// TIA Portal project "DnomaidDBMS" (V13) (continued)
REGION Network 8: dA..Data Select
         L     #Network_8;
         T     #P_RET_VAL.MEM;
         A(;
         L     #COUNT.dA00;
         L     0;
         <>I;
         );
         A(;
         L     #COUNT.dA00;
         L     #QuantityDB;
         <=I;
         );
         JC    dA00;
         L     1;
         T     #COUNT.dA00;
         JU    dA00;
   dA00: NOP   0;
         L     #COUNT.dA00;
         JL    dAXX;
         JU    dAXX;
         JU    dA11;  //db[1]
         JU    dA21;  //db[2]
         JU    dA31;  //db[3]
         JU    dA41;  //db[4]
         JU    dA51;  //db[5]
         JU    dA61;  //db[6]
   dAXX: JU    dZFF;  //end
   dA11: NOP   0;
         L     #COUNT.dA00;
         T     #Status.Mem.SelctBBDDNum;
         SET;
         R     #AUX.FullDatabase;
         A     #Status.Perm.Push_nDB[1];
         AN    #Status.Mem.Full_nDB[1];
         =     #AUX.PushDatabase;
         JCN   dA12;
         L     #P_RET_VAL.MEM;
         T     #P_RET_VAL.V[1];
         T     #P_RET_VAL.V[2];
         CALL  FILL
         ( BVAL    := #ANY_DB1_FE,
           RET_VAL := #P_RET_VAL.V[1],
           BLK     := #ANY_DB1_IE
         );
         L     #P_RET_VAL.V[1];
         L     0;
         <>I;
         S     #FAULT;
         JC    END;
         CALL  FILL
         ( BVAL    := #IniData,
           RET_VAL := #P_RET_VAL.V[2],
           BLK     := #ANY_DB1_F
         );
         L     #P_RET_VAL.V[2];
         L     0;
         <>I;
         S     #FAULT;
         JC    END;
         R     #Status.Perm.Push_nDB[1];
         JU    dWFF;
   dA12: NOP   0;
         OPN   DB[ #LIST_DB_T.DbNumber[1]];
         LAR1  #""Address_104";
         L     LD[AR1, P#0.0];
         T     #AUX.LD_01;
         L     LW[AR1, P#4.0];
         T     #AUX.LW_01;
         L     LD[AR1, P#6.0];
         T     #AUX.LD_02;
         LAR1  #""Address_290";  //SEL
         L     #AUX.LD_01;
         T     LD[AR1, P#0.0];
         L     #AUX.LW_01;
         T     LW[AR1, P#4.0];
         L     #AUX.LD_02;
         T     LD[AR1, P#6.0];
         T     #P_ADR.I;
         LAR1  #""Address_113";
         L     LD[AR1, P#0.0];
         T     #AUX.LD_01;
         L     LW[AR1, P#4.0];
         T     #AUX.LW_01;
         L     LD[AR1, P#6.0];
         T     #AUX.LD_02;
         LAR1  #""Address_293";  //SEL
         L     #AUX.LD_01;
         T     LD[AR1, P#0.0];
         L     #AUX.LW_01;
         T     LW[AR1, P#4.0];
         L     #AUX.LD_02;
         T     LD[AR1, P#6.0];
         T     #P_ADR.F;
         JU    dAFF;
   dA21: NOP   0;
         L     #COUNT.dA00;
         T     #Status.Mem.SelctBBDDNum;
         SET;
         R     #AUX.FullDatabase;
         A     #Status.Perm.Push_nDB[2];
         AN    #Status.Mem.Full_nDB[2];
         =     #AUX.PushDatabase;
         JCN   dA22;
         L     #P_RET_VAL.MEM;
         T     #P_RET_VAL.V[1];
         T     #P_RET_VAL.V[2];
         CALL  FILL
         ( BVAL    := #ANY_DB2_FE,
           RET_VAL := #P_RET_VAL.V[1],
           BLK     := #ANY_DB2_IE
         );
         L     #P_RET_VAL.V[1];
         L     0;
         <>I;
         S     #FAULT;
         JC    END;
         CALL  FILL
         ( BVAL    := #IniData,
           RET_VAL := #P_RET_VAL.V[2],
           BLK     := #ANY_DB2_F
         );
         L     #P_RET_VAL.V[2];
         L     0;
         <>I;
         S     #FAULT;
         JC    END;
         R     #Status.Perm.Push_nDB[2];
         JU    dWFF;
   dA22: NOP   0;
         OPN   DB[ #LIST_DB_T.DbNumber[2]];
         LAR1  #""Address_119";
         L     LD[AR1, P#0.0];
         T     #AUX.LD_01;
         L     LW[AR1, P#4.0];
         T     #AUX.LW_01;
         L     LD[AR1, P#6.0];
         T     #AUX.LD_02;
         LAR1  #""Address_290";  //SEL
         L     #AUX.LD_01;
         T     LD[AR1, P#0.0];
         L     #AUX.LW_01;
         T     LW[AR1, P#4.0];
         L     #AUX.LD_02;
         T     LD[AR1, P#6.0];
         T     #P_ADR.I;
         LAR1  #""Address_126";
         L     LD[AR1, P#0.0];
         T     #AUX.LD_01;
         L     LW[AR1, P#4.0];
         T     #AUX.LW_01;
         L     LD[AR1, P#6.0];
         T     #AUX.LD_02;
         LAR1  #""Address_293";  //SELECT
         L     #AUX.LD_01;
         T     LD[AR1, P#0.0];
         L     #AUX.LW_01;
         T     LW[AR1, P#4.0];
         L     #AUX.LD_02;
         T     LD[AR1, P#6.0];
         T     #P_ADR.F;
         JU    dAFF;
   dA31: NOP   0;
         L     #COUNT.dA00;
         T     #Status.Mem.SelctBBDDNum;
         SET;
         R     #AUX.FullDatabase;
         A     #Status.Perm.Push_nDB[3];
         AN    #Status.Mem.Full_nDB[3];
         =     #AUX.PushDatabase;
         JCN   dA32;
         L     #P_RET_VAL.MEM;
         T     #P_RET_VAL.V[1];
         T     #P_RET_VAL.V[2];
         CALL  FILL
         ( BVAL    := #ANY_DB3_FE,
           RET_VAL := #P_RET_VAL.V[1],
           BLK     := #ANY_DB3_IE
         );
         L     #P_RET_VAL.V[1];
         L     0;
         <>I;
         S     #FAULT;
         JC    END;
         CALL  FILL
         ( BVAL    := #IniData,
           RET_VAL := #P_RET_VAL.V[2],
           BLK     := #ANY_DB3_F
         );
         L     #P_RET_VAL.V[2];
         L     0;
         <>I;
         S     #FAULT;
         JC    END;
         R     #Status.Perm.Push_nDB[3];
         JU    dWFF;
   dA32: NOP   0;
         OPN   DB[ #LIST_DB_T.DbNumber[3]];
         LAR1  #""Address_132";
         L     LD[AR1, P#0.0];
         T     #AUX.LD_01;
         L     LW[AR1, P#4.0];
         T     #AUX.LW_01;
         L     LD[AR1, P#6.0];
         T     #AUX.LD_02;
         LAR1  #""Address_290";  //SEL
         L     #AUX.LD_01;
         T     LD[AR1, P#0.0];
         L     #AUX.LW_01;
         T     LW[AR1, P#4.0];
         L     #AUX.LD_02;
         T     LD[AR1, P#6.0];
         T     #P_ADR.I;
         LAR1  #""Address_139";
         L     LD[AR1, P#0.0];
         T     #AUX.LD_01;
         L     LW[AR1, P#4.0];
         T     #AUX.LW_01;
         L     LD[AR1, P#6.0];
         T     #AUX.LD_02;
         LAR1  #""Address_293";  //SEL
         L     #AUX.LD_01;
         T     LD[AR1, P#0.0];
         L     #AUX.LW_01;
         T     LW[AR1, P#4.0];
         L     #AUX.LD_02;
         T     LD[AR1, P#6.0];
         T     #P_ADR.F;
         JU    dAFF;
   dA41: NOP   0;
         L     #COUNT.dA00;
         T     #Status.Mem.SelctBBDDNum;
         SET;
         R     #AUX.FullDatabase;
         A     #Status.Perm.Push_nDB[4];
         AN    #Status.Mem.Full_nDB[4];
         =     #AUX.PushDatabase;
         JCN   dA42;
         L     #P_RET_VAL.MEM;
         T     #P_RET_VAL.V[1];
         T     #P_RET_VAL.V[2];
         CALL  FILL
         ( BVAL    := #ANY_DB4_FE,
           RET_VAL := #P_RET_VAL.V[1],
           BLK     := #ANY_DB4_IE
         );
         L     #P_RET_VAL.V[1];
         L     0;
         <>I;
         S     #FAULT;
         JC    END;
         CALL  FILL
         ( BVAL    := #IniData,
           RET_VAL := #P_RET_VAL.V[2],
           BLK     := #ANY_DB4_F
         );
         L     #P_RET_VAL.V[2];
         L     0;
         <>I;
         S     #FAULT;
         JC    END;
         R     #Status.Perm.Push_nDB[4];
         JU    dWFF;
   dA42: NOP   0;
         OPN   DB[ #LIST_DB_T.DbNumber[4]];
         LAR1  #""Address_145";
         L     LD[AR1, P#0.0];
         T     #AUX.LD_01;
         L     LW[AR1, P#4.0];
         T     #AUX.LW_01;
         L     LD[AR1, P#6.0];
         T     #AUX.LD_02;
         LAR1  #""Address_290";  //SEL
         L     #AUX.LD_01;
         T     LD[AR1, P#0.0];
         L     #AUX.LW_01;
         T     LW[AR1, P#4.0];
         L     #AUX.LD_02;
         T     LD[AR1, P#6.0];
         T     #P_ADR.I;
         LAR1  #""Address_152";
         L     LD[AR1, P#0.0];
         T     #AUX.LD_01;
         L     LW[AR1, P#4.0];
         T     #AUX.LW_01;
         L     LD[AR1, P#6.0];
         T     #AUX.LD_02;
         LAR1  #""Address_293";  //SEL
         L     #AUX.LD_01;
         T     LD[AR1, P#0.0];
         L     #AUX.LW_01;
         T     LW[AR1, P#4.0];
         L     #AUX.LD_02;
         T     LD[AR1, P#6.0];
         T     #P_ADR.F;
         JU    dAFF;
   dA51: NOP   0;
         L     #COUNT.dA00;
         T     #Status.Mem.SelctBBDDNum;
         SET;
         R     #AUX.FullDatabase;
         A     #Status.Perm.Push_nDB[5];
         AN    #Status.Mem.Full_nDB[5];
         =     #AUX.PushDatabase;
         JCN   dA52;
         L     #P_RET_VAL.MEM;
         T     #P_RET_VAL.V[1];
         T     #P_RET_VAL.V[2];
         CALL  FILL
         ( BVAL    := #ANY_DB5_FE,
           RET_VAL := #P_RET_VAL.V[1],
           BLK     := #ANY_DB5_IE
         );
         L     #P_RET_VAL.V[1];
         L     0;
         <>I;
         S     #FAULT;
         JC    END;
         CALL  FILL
         ( BVAL    := #IniData,
           RET_VAL := #P_RET_VAL.V[2],
           BLK     := #ANY_DB5_F
         );
         L     #P_RET_VAL.V[2];
         L     0;
         <>I;
         S     #FAULT;
         JC    END;
         R     #Status.Perm.Push_nDB[5];
         JU    dWFF;
   dA52: NOP   0;
         OPN   DB[ #LIST_DB_T.DbNumber[5]];
         LAR1  #""Address_158";
         L     LD[AR1, P#0.0];
         T     #AUX.LD_01;
         L     LW[AR1, P#4.0];
         T     #AUX.LW_01;
         L     LD[AR1, P#6.0];
         T     #AUX.LD_02;
         LAR1  #""Address_290";  //SEL
         L     #AUX.LD_01;
         T     LD[AR1, P#0.0];
         L     #AUX.LW_01;
         T     LW[AR1, P#4.0];
         L     #AUX.LD_02;
         T     LD[AR1, P#6.0];
         T     #P_ADR.I;
         LAR1  #""Address_165";
         L     LD[AR1, P#0.0];
         T     #AUX.LD_01;
         L     LW[AR1, P#4.0];
         T     #AUX.LW_01;
         L     LD[AR1, P#6.0];
         T     #AUX.LD_02;
         LAR1  #""Address_293";  //SEL
         L     #AUX.LD_01;
         T     LD[AR1, P#0.0];
         L     #AUX.LW_01;
         T     LW[AR1, P#4.0];
         L     #AUX.LD_02;
         T     LD[AR1, P#6.0];
         T     #P_ADR.F;
         JU    dAFF;
   dA61: NOP   0;
         L     #COUNT.dA00;
         T     #Status.Mem.SelctBBDDNum;
         SET;
         R     #AUX.FullDatabase;
         A     #Status.Perm.Push_nDB[6];
         AN    #Status.Mem.Full_nDB[6];
         =     #AUX.PushDatabase;
         JCN   dA62;
         L     #P_RET_VAL.MEM;
         T     #P_RET_VAL.V[1];
         T     #P_RET_VAL.V[2];
         CALL  FILL
         ( BVAL    := #ANY_DB6_FE,
           RET_VAL := #P_RET_VAL.V[1],
           BLK     := #ANY_DB6_IE
         );
         L     #P_RET_VAL.V[1];
         L     0;
         <>I;
         S     #FAULT;
         JC    END;
         CALL  FILL
         ( BVAL    := #IniData,
           RET_VAL := #P_RET_VAL.V[2],
           BLK     := #ANY_DB6_F
         );
         L     #P_RET_VAL.V[2];
         L     0;
         <>I;
         S     #FAULT;
         JC    END;
         R     #Status.Perm.Push_nDB[6];
         JU    dWFF;
   dA62: NOP   0;
         OPN   DB[ #LIST_DB_T.DbNumber[6]];
         LAR1  #""Address_171";
         L     LD[AR1, P#0.0];
         T     #AUX.LD_01;
         L     LW[AR1, P#4.0];
         T     #AUX.LW_01;
         L     LD[AR1, P#6.0];
         T     #AUX.LD_02;
         LAR1  #""Address_290";  //SEL
         L     #AUX.LD_01;
         T     LD[AR1, P#0.0];
         L     #AUX.LW_01;
         T     LW[AR1, P#4.0];
         L     #AUX.LD_02;
         T     LD[AR1, P#6.0];
         T     #P_ADR.I;
         LAR1  #""Address_178";
         L     LD[AR1, P#0.0];
         T     #AUX.LD_01;
         L     LW[AR1, P#4.0];
         T     #AUX.LW_01;
         L     LD[AR1, P#6.0];
         T     #AUX.LD_02;
         LAR1  #""Address_293";  //SEL
         L     #AUX.LD_01;
         T     LD[AR1, P#0.0];
         L     #AUX.LW_01;
         T     LW[AR1, P#4.0];
         L     #AUX.LD_02;
         T     LD[AR1, P#6.0];
         T     #P_ADR.F;
         JU    dAFF;
   dAFF: NOP   0;
END_REGION

REGION Network 9: dC..Data Search empty space
         LAR1  #P_ADR.I;
         JU    dC00;
   dC00: NOP   0;
         L     #Network_9;
         T     #P_RET_VAL.MEM;
         TAR1;
         T     #SAVE_AR1.dC00;
         L     1;
   dC01: NOP   0;
         T     #COUNT.dC00;
         L     DBB[AR1, P#0.0];
         L     ' ';
         <>I;
         =     #AUX.DifferentValue;
         AN    #AUX.DifferentValue;
         JC    dCFF;
         L     #P_ADR.F;
         L     #SAVE_AR1.dC00;
         <=D;
         =     #AUX.FullDatabase;
         A     #AUX.FullDatabase;
         JC    dCWF;
         L     P#1.0;
         +AR1;
         L     #COUNT.dC00;
         LOOP  dC01;
         L     #SAVE_AR1.dC00;
         LAR1;
         L     #LENGTH.PointerData;
         +AR1;
         JU    dC00;
END_REGION

REGION Network 10: dC..Data Full
         JU    dCWF;
   dCWF: NOP   0;
         L     #Network_10;
         T     #P_RET_VAL.MEM;
         AN    #AUX.FullDatabase;
         JC    dCWW;
         L     #Status.Mem.SelctBBDDNum;
         JL    dCXX;
         JU    dCEE;  //fault
         JU    dC11;  //db[1]
         JU    dC12;  //db[2]
         JU    dC13;  //db[3]
         JU    dC14;  //db[4]
         JU    dC15;  //db[5]
         JU    dC16;  //db[6]
   dCXX: JU    dCEE;  //fault
   dC11: NOP   0;
         A     #AUX.FullDatabase;
         =     #Status.Mem.Full_nDB[1];
         JU    dCWW;
   dC12: NOP   0;
         A     #AUX.FullDatabase;
         =     #Status.Mem.Full_nDB[2];
         JU    dCWW;
   dC13: NOP   0;
         A     #AUX.FullDatabase;
         =     #Status.Mem.Full_nDB[3];
         JU    dCWW;
   dC14: NOP   0;
         A     #AUX.FullDatabase;
         =     #Status.Mem.Full_nDB[4];
         JU    dCWW;
   dC15: NOP   0;
         A     #AUX.FullDatabase;
         =     #Status.Mem.Full_nDB[5];
         JU    dCWW;
   dC16: NOP   0;
         A     #AUX.FullDatabase;
         =     #Status.Mem.Full_nDB[6];
         JU    dCWW;
   dCEE: NOP   0;
         SET;
         S     #FAULT;
         JU    END;
   dCWW: NOP   0;
         JU    dWFF;
         JU    dCFF;
   dCFF: NOP   0;
END_REGION

REGION Network 11: dD..Data Find space
         JU    dD00;
   dD00: NOP   0;
         L     #Network_11;
         T     #P_RET_VAL.MEM;
         L     #SAVE_AR1.dC00;
         LAR1;
         L     #LENGTH.PointerData;
         +AR1;
         L     #P_ADR.F;
         TAR1;
         <D;
         JC    dWFF;
         JU    dDFF;
   dDFF: NOP   0;
END_REGION

REGION Network 12: dE..Data Find data
         JU    dE00;
   dE00: NOP   0;
         L     #Network_12;
         T     #P_RET_VAL.MEM;
         TAR1;
         T     #SAVE_AR1.dE00;
         L     1;
   dE01: NOP   0;
         T     #COUNT.dE00;
         L     DBB[AR1, P#0.0];
         L     ' ';
         ==I;
         =     #AUX.EmptyData;
         AN    #AUX.EmptyData;
         JC    dEFF;
         L     #P_ADR.F;
         L     #SAVE_AR1.dE00;
         <=D;
         JC    dWFF;
         L     P#1.0;
         +AR1;
         L     #COUNT.dE00;
         LOOP  dE01;
         L     #SAVE_AR1.dE00;
         LAR1;
         L     #LENGTH.PointerData;
         +AR1;
         JU    dE00;
         JU    dEFF;
   dEFF: NOP   0;
END_REGION

REGION Network 13: dF..Data Move data
         JU    dF01;
   dF01: NOP   0;
         L     #Network_13;
         T     #P_RET_VAL.MEM;
         L     #SAVE_AR1.dE00;
         T     #P_ADR.F;
         LAR1  #""Address_293";
         T     LD[AR1, P#6.0];
         L     #SAVE_AR1.dC00;
         T     #P_ADR.I;
         LAR1  #""Address_290";
         T     LD[AR1, P#6.0];
         LAR1;
         L     #P_RET_VAL.MEM;
         T     #P_RET_VAL.V[1];
         T     #P_RET_VAL.V[2];
         CALL  FILL
         ( BVAL    := #ANY_DB_SELECT_F,
           RET_VAL := #P_RET_VAL.V[1],
           BLK     := #ANY_DB_SELECT_I
         );
         L     #P_RET_VAL.V[1];
         L     0;
         <>I;
         S     #FAULT;
         JC    END;
         CALL  FILL
         ( BVAL    := #IniData,
           RET_VAL := #P_RET_VAL.V[2],
           BLK     := #ANY_DB_SELECT_F
         );
         L     #P_RET_VAL.V[2];
         L     0;
         <>I;
         S     #FAULT;
         JC    END;
         JU    dZFF;
   dWFF: NOP   0;
         L     #COUNT.dA00;
         +     1;
         T     #COUNT.dA00;
         L     #QuantityDB;
         >I;
         JC    dZFF;
         JU    dA00;
   //--->END
         JU    dZFF;
   dZFF: NOP   0;
END_REGION

REGION Network 14: fA..Query
         JU    fA0X;
   fA0X: NOP   0;
         L     #Network_14;
         T     #P_RET_VAL.MEM;
         AN    #Request.Query.Request;
         R     #Response.Query.DataAvailable;
         R     #Response.Query.DataNotAvailable;
         NOT;
         FP    #FP_REQUEST.QueryDB;
         JC    fA0Y;
         JU    fBFF;
   fA0Y: NOP   0;
         L     #P_RET_VAL.MEM;
         T     #P_RET_VAL.V[1];
         T     #P_RET_VAL.V[2];
         CALL  FILL
         ( BVAL    := #Request.Query.BarcodeDig,
           RET_VAL := #P_RET_VAL.V[1],
           BLK     := #DigitFilter
         );
         L     #P_RET_VAL.V[1];
         L     0;
         <>I;
         S     #FAULT;
         JC    END;
         JU    jA00;  //Goto Data input filters
   fAR2: NOP   0;  //Return Data input filters
         CALL  FILL
         ( BVAL    := #DigitFilter,
           RET_VAL := #P_RET_VAL.V[2],
           BLK     := #QueryData
         );
         L     #P_RET_VAL.V[2];
         L     0;
         <>I;
         S     #FAULT;
         JC    END;
         CALL  FILL
         ( BVAL    := #IniData,
           RET_VAL := #P_RET_VAL.V[3],
           BLK     := #Response.QueryDataAvailable
         );
         L     #P_RET_VAL.V[3];
         L     0;
         <>I;
         S     #FAULT;
         JC    END;
         AN    #DataInputOK;
         JC    fB50;  //Error data input
         L     1;
         T     #COUNT.fA00;
   fA00: NOP   0;
         L     #COUNT.fA00;
         JL    fAXX;
         JU    fAXX;
         JU    fA11;  //db[1]
         JU    fA21;  //db[2]
         JU    fA31;  //db[3]
         JU    fA41;  //db[4]
         JU    fA51;  //db[5]
         JU    fA61;  //db[6]
         JU    fB40;  //end
   fAXX: JU    fAEE;  //fault
   fA11: NOP   0;
         OPN   DB[ #LIST_DB_T.DbNumber[1]];
         LAR1  #P_ADR.I_DB[1];
         L     #NumDataArrayDB[1];
         JU    fA10;
   fA21: NOP   0;
         OPN   DB[ #LIST_DB_T.DbNumber[2]];
         LAR1  #P_ADR.I_DB[2];
         L     #NumDataArrayDB[2];
         JU    fA10;
   fA31: NOP   0;
         OPN   DB[ #LIST_DB_T.DbNumber[3]];
         LAR1  #P_ADR.I_DB[3];
         L     #NumDataArrayDB[3];
         JU    fA10;
   fA41: NOP   0;
         OPN   DB[ #LIST_DB_T.DbNumber[4]];
         LAR1  #P_ADR.I_DB[4];
         L     #NumDataArrayDB[4];
         JU    fA10;
   fA51: NOP   0;
         OPN   DB[ #LIST_DB_T.DbNumber[5]];
         LAR1  #P_ADR.I_DB[5];
         L     #NumDataArrayDB[5];
         JU    fA10;
   fA61: NOP   0;
         OPN   DB[ #LIST_DB_T.DbNumber[6]];
         LAR1  #P_ADR.I_DB[6];
         L     #NumDataArrayDB[6];
         JU    fA10;
   fA10: NOP   0;
         T     #COUNT.fA01;
         TAR1;
         T     #SAVE_AR1.fA10;
         SET;
   //-------------------------------
         TAR1;
         T     #P_ADR.SAVE_COMP_01;
         T     #P_ADR.COMP_01;
         L     #""Address_347";
         T     #P_ADR.COMP_02;
         SET;
         R     #AUX.DifferentValue;
         L     #LENGTH.Code;
   fMP0: NOP   0;
         T     #COUNT.fA02;
         LAR1  #P_ADR.COMP_01;
         L     DBB[AR1, P#0.0];
         LAR1  #P_ADR.COMP_02;
         L     DIB[AR1, P#0.0];
         <>I;
         S     #AUX.DifferentValue;
         L     P#1.0;
         L     #P_ADR.COMP_01;
         +D;
         T     #P_ADR.COMP_01;
         L     P#1.0;
         L     #P_ADR.COMP_02;
         +D;
         T     #P_ADR.COMP_02;
         L     #COUNT.fA02;
         LOOP  fMP0;
         LAR1  #P_ADR.SAVE_COMP_01;
   //-------------------------------
         AN    #AUX.DifferentValue;
         JC    fB20;
         L     #LENGTH.PointerData;
         +AR1;
         L     #COUNT.fA01;
         LOOP  fA10;
         JU    fWFF;
   fWFF: NOP   0;
         L     #COUNT.fA00;
         +     1;
         T     #COUNT.fA00;
         L     #QuantityDB;
         >I;
         JC    fB40;
         JU    fA00;
   fAEE: NOP   0;
         SET;
         S     #FAULT;
         JU    END;
         JU    fAFF;
   fAFF: NOP   0;
         JU    END;
   fB20: NOP   0;
         L     #COUNT.fA00;
         JL    fB3X;
         JU    fB3X;
         JU    fB31;  //db[1]
         JU    fB32;  //db[2]
         JU    fB33;  //db[3]
         JU    fB34;  //db[4]
         JU    fB35;  //db[5]
         JU    fB36;  //db[6]
   fB3X: JU    fB3E;  //fault
   fB31: NOP   0;
         LAR1  #""Address_104";
         JU    fB3F;
   fB32: NOP   0;
         LAR1  #""Address_119";
         JU    fB3F;
   fB33: NOP   0;
         LAR1  #""Address_132";
         JU    fB3F;
   fB34: NOP   0;
         LAR1  #""Address_145";
         JU    fB3F;
   fB35: NOP   0;
         LAR1  #""Address_158";
         JU    fB3F;
   fB36: NOP   0;
         LAR1  #""Address_171";
         JU    fB3F;
   fB3E: NOP   0;
         SET;
         S     #FAULT;
         JU    END;
         JU    fB3F;
   fB3F: NOP   0;
         L     LD[AR1, P#0.0];
         T     #AUX.LD_01;
         L     LW[AR1, P#4.0];
         T     #AUX.LW_01;
         T     #PAUXnDB;
         LAR1  #""Address_381";
         L     #AUX.LD_01;
         T     LD[AR1, P#0.0];
         L     #AUX.LW_01;
         T     LW[AR1, P#4.0];
         L     #SAVE_AR1.fA10;
         T     LD[AR1, P#6.0];
         L     #P_RET_VAL.MEM;
         T     #P_RET_VAL.V[1];
         CALL  FILL
         ( BVAL    := #ANY_DB_QUERY,
           RET_VAL := #P_RET_VAL.V[1],
           BLK     := #Response.QueryDataAvailable
         );
         L     #P_RET_VAL.V[1];
         L     0;
         <>I;
         S     #FAULT;
         JC    END;
         S     #Response.Query.DataAvailable;
         R     #Response.Query.DataNotAvailable;
         L     #LogDataAvailable;
         T     #Log.Request;
         JU    fB50;
   fB40: NOP   0;
         SET;
         R     #Response.Query.DataAvailable;
         S     #Response.Query.DataNotAvailable;
         L     #LogDataNotAvailable;
         T     #Log.Request;
   fB50: NOP   0;
         A     #DataInputOK;
         JC    fB51;  //Error data input
         L     #LogDataInputNOK;
         T     #Log.Request;
   fB51: NOP   0;
         L     #P_RET_VAL.MEM;
         T     #P_RET_VAL.V[1];
         CALL  FILL
         ( BVAL    := #QueryData,
           RET_VAL := #P_RET_VAL.V[1],
           BLK     := #Response.Query.BarcodeDig
         );
         L     #P_RET_VAL.V[1];
         L     0;
         <>I;
         S     #FAULT;
         JC    END;
         CALL  FILL
         ( BVAL    := #QueryData,
           RET_VAL := #P_RET_VAL.V[2],
           BLK     := #Log.DatabaseTable
         );
         L     #P_RET_VAL.V[2];
         L     0;
         <>I;
         S     #FAULT;
         JC    END;
         CALL  FILL
         ( BVAL    := #DateTime,
           RET_VAL := #P_RET_VAL.V[3],
           BLK     := #Log.DatabaseTable.DateTime
         );
         L     #P_RET_VAL.V[3];
         L     0;
         <>I;
         S     #FAULT;
         JC    END;
         JU    fBFF;
   fBFF: NOP   0;
END_REGION

REGION Network 15: gA..Insert
         JU    gA00;
   gA00: NOP   0;
         L     #Network_15;
         T     #P_RET_VAL.MEM;
         SET;
   //      R     #AUX.StatusPermInsert_nDB
         AN    #Request.Insert.Request;
         R     #Response.Insert.Completed;
         L     #QuantityDB;
         T     #COUNT.gA00;
         NOP   0;
         SET;
         L     #COUNT.gA00;
         JL    gAXX;
         JU    gAXX;
         JU    gA11;  //db[1]
         JU    gA21;  //db[2]
         JU    gA31;  //db[3]
         JU    gA41;  //db[4]
         JU    gA51;  //db[5]
         JU    gA61;  //db[6]
   gAXX: JU    gAEE;  //fault
   gA11: NOP   0;
         A     #Status.Perm.Insert_nDB[1];
         JU    gA01;
   gA21: NOP   0;
         A     #Status.Perm.Insert_nDB[2];
         JU    gA01;
   gA31: NOP   0;
         A     #Status.Perm.Insert_nDB[3];
         JU    gA01;
   gA41: NOP   0;
         A     #Status.Perm.Insert_nDB[4];
         JU    gA01;
   gA51: NOP   0;
         A     #Status.Perm.Insert_nDB[5];
         JU    gA01;
   gA61: NOP   0;
         A     #Status.Perm.Insert_nDB[6];
         JU    gA01;
   gAEE: NOP   0;
         SET;
         S     #FAULT;
         JU    END;
   gA01: NOP   0;
         =     #AUX.StatusPermInsert_nDB;
         A     #AUX.TON_StatusPermInsert_nDB;
         AN    #Status.Mem.FillAll;
         AN    #Status.Fb_Fault;
         =     #Status.Perm.Insert;
         A     #FULL;  //Data base full
         JC    gA02;
         A     #Request.Query.Request;
         JC    gAFF;
         A     #AUX.TON_StatusPermInsert_nDB;
   gA02: NOP   0;
         A     #Request.Insert.Request;
         FP    #FP_REQUEST.InsertDB;
         JC    gA03;
         JU    gAFF;
   gA03: NOP   0;
         L     #P_RET_VAL.MEM;
         T     #P_RET_VAL.V[1];
         T     #P_RET_VAL.V[2];
         T     #P_RET_VAL.V[3];
         T     #P_RET_VAL.V[4];
         T     #P_RET_VAL.V[5];
         CALL  FILL
         ( BVAL    := #Request.Insert.BarcodeData,
           RET_VAL := #P_RET_VAL.V[1],
           BLK     := #DigitFilter
         );
         L     #P_RET_VAL.V[1];
         L     0;
         <>I;
         S     #FAULT;
         JC    END;
         JU    jA00;  //Goto Data input filters
   gAR2: NOP   0;  //Return Data input filters
         CALL  FILL
         ( BVAL    := #DigitFilter,
           RET_VAL := #P_RET_VAL.V[2],
           BLK     := #InsertData.BarcodeData
         );
         L     #P_RET_VAL.V[2];
         L     0;
         <>I;
         S     #FAULT;
         JC    END;
         CALL  FILL
         ( BVAL    := #DateTime,
           RET_VAL := #P_RET_VAL.V[3],
           BLK     := #InsertData.DateTime
         );
         L     #P_RET_VAL.V[3];
         L     0;
         <>I;
         S     #FAULT;
         JC    END;
         AN    #DataInputOK;
         S     #DATA_ERROR;
         JC    gA05;  //Error data input
         A     #FULL;
         S     #DATA_ERROR;
         JC    gA06;  //Data base full
         L     #COUNT.gA00;
         JL    gBXX;
         JU    gBXX;
         JU    gB11;  //db[1]
         JU    gB21;  //db[2]
         JU    gB31;  //db[3]
         JU    gB41;  //db[4]
         JU    gB51;  //db[5]
         JU    gB61;  //db[6]
   gBXX: JU    gBEE;  //fault
   gB11: NOP   0;
         CALL  FILL
         ( BVAL    := #InsertData,
           RET_VAL := #P_RET_VAL.V[3],
           BLK     := #ANY_DB1_F
         );
         L     #P_RET_VAL.V[3];
         L     0;
         <>I;
         S     #FAULT;
         JC    END;
         JU    gA04;
   gB21: NOP   0;
         CALL  FILL
         ( BVAL    := #InsertData,
           RET_VAL := #P_RET_VAL.V[3],
           BLK     := #ANY_DB2_F
         );
         L     #P_RET_VAL.V[3];
         L     0;
         <>I;
         S     #FAULT;
         JC    END;
         JU    gA04;
   gB31: NOP   0;
         CALL  FILL
         ( BVAL    := #InsertData,
           RET_VAL := #P_RET_VAL.V[3],
           BLK     := #ANY_DB3_F
         );
         L     #P_RET_VAL.V[3];
         L     0;
         <>I;
         S     #FAULT;
         JC    END;
         JU    gA04;
   gB41: NOP   0;
         CALL  FILL
         ( BVAL    := #InsertData,
           RET_VAL := #P_RET_VAL.V[3],
           BLK     := #ANY_DB4_F
         );
         L     #P_RET_VAL.V[3];
         L     0;
         <>I;
         S     #FAULT;
         JC    END;
         JU    gA04;
   gB51: NOP   0;
         CALL  FILL
         ( BVAL    := #InsertData,
           RET_VAL := #P_RET_VAL.V[3],
           BLK     := #ANY_DB5_F
         );
         L     #P_RET_VAL.V[3];
         L     0;
         <>I;
         S     #FAULT;
         JC    END;
         JU    gA04;
   gB61: NOP   0;
         CALL  FILL
         ( BVAL    := #InsertData,
           RET_VAL := #P_RET_VAL.V[3],
           BLK     := #ANY_DB6_F
         );
         L     #P_RET_VAL.V[3];
         L     0;
         <>I;
         S     #FAULT;
         JC    END;
         JU    gA04;
   gBEE: NOP   0;
         SET;
         S     #FAULT;
         JU    END;
   gA04: NOP   0;
         CALL  FILL
         ( BVAL    := #InsertData,
           RET_VAL := #P_RET_VAL.V[4],
           BLK     := #Response.InsertData
         );
         L     #P_RET_VAL.V[4];
         L     0;
         <>I;
         S     #FAULT;
         JC    END;
         S     #Response.Insert.Completed;
         L     #LogInsert;
         T     #Log.Request;
         A     #DataInputOK;
         JC    gA07;
   gA05: NOP   0;
         L     #LogDataInputNOK;  //Data input NOK
         T     #Log.Request;
         SET;
         JU    gA07;
   gA06: NOP   0;
         L     #LogFullData;  //Data base full
         T     #Log.Request;
         SET;
         JU    gA07;
   gA07: NOP   0;
         CALL  FILL
         ( BVAL    := #InsertData,
           RET_VAL := #P_RET_VAL.V[5],
           BLK     := #Log.DatabaseTable
         );
         L     #P_RET_VAL.V[5];
         L     0;
         <>I;
         S     #FAULT;
         JC    END;
         JU    gAFF;
   gAFF: NOP   0;
END_REGION

REGION Network 16: hA..Delete
         JU    hA0X;
   hA0X: NOP   0;
         L     #Network_16;
         T     #P_RET_VAL.MEM;
         AN    #Request.Delete.Request;
         R     #Response.Delete.Completed;
         NOT;
         FP    #FP_REQUEST.DeleteDB;
         JC    hA0Y;
         JU    hBFF;
   hA0Y: NOP   0;
         L     #P_RET_VAL.MEM;
         T     #P_RET_VAL.V[1];
         T     #P_RET_VAL.V[2];
         CALL  FILL
         ( BVAL    := #Request.Delete.BarcodeDig,
           RET_VAL := #P_RET_VAL.V[1],
           BLK     := #DigitFilter
         );
         L     #P_RET_VAL.V[1];
         L     0;
         <>I;
         S     #FAULT;
         JC    END;
         JU    jA00;  //Goto Data input filters
   hAR2: NOP   0;  //Return Data input filters
         CALL  FILL
         ( BVAL    := #DigitFilter,
           RET_VAL := #P_RET_VAL.V[2],
           BLK     := #DeleteData
         );
         L     #P_RET_VAL.V[2];
         L     0;
         <>I;
         S     #FAULT;
         JC    END;
         CALL  FILL
         ( BVAL    := #IniData,
           RET_VAL := #P_RET_VAL.V[3],
           BLK     := #Response.DeleteData
         );
         L     #P_RET_VAL.V[3];
         L     0;
         <>I;
         S     #FAULT;
         AN    #DataInputOK;
         JC    hB3G;  //Error data input
         L     1;
         T     #COUNT.hA00;
   hA00: NOP   0;
         L     #COUNT.hA00;
         JL    hAXX;
         JU    hAXX;
         JU    hA11;  //db[1]
         JU    hA21;  //db[2]
         JU    hA31;  //db[3]
         JU    hA41;  //db[4]
         JU    hA51;  //db[5]
         JU    hA61;  //db[6]
         JU    hB40;  //end
   hAXX: JU    hAEE;  //fault
   hA11: NOP   0;
         OPN   DB[ #LIST_DB_T.DbNumber[1]];
         LAR1  #P_ADR.I_DB[1];
         L     #NumDataArrayDB[1];
         JU    hA10;
   hA21: NOP   0;
         OPN   DB[ #LIST_DB_T.DbNumber[2]];
         LAR1  #P_ADR.I_DB[2];
         L     #NumDataArrayDB[2];
         JU    hA10;
   hA31: NOP   0;
         OPN   DB[ #LIST_DB_T.DbNumber[3]];
         LAR1  #P_ADR.I_DB[3];
         L     #NumDataArrayDB[3];
         JU    hA10;
   hA41: NOP   0;
         OPN   DB[ #LIST_DB_T.DbNumber[4]];
         LAR1  #P_ADR.I_DB[4];
         L     #NumDataArrayDB[4];
         JU    hA10;
   hA51: NOP   0;
         OPN   DB[ #LIST_DB_T.DbNumber[5]];
         LAR1  #P_ADR.I_DB[5];
         L     #NumDataArrayDB[5];
         JU    hA10;
   hA61: NOP   0;
         OPN   DB[ #LIST_DB_T.DbNumber[6]];
         LAR1  #P_ADR.I_DB[6];
         L     #NumDataArrayDB[6];
         JU    hA10;
   hA10: NOP   0;
         T     #COUNT.hA01;
         TAR1;
         T     #SAVE_AR1.hA10;
         SET;
   //-------------------------------
         TAR1;
         T     #P_ADR.SAVE_COMP_01;
         T     #P_ADR.COMP_01;
         L     #""Address_433";
         T     #P_ADR.COMP_02;
         SET;
         R     #AUX.DifferentValue;
         L     #LENGTH.Code;
   hMP0: NOP   0;
         T     #COUNT.hA02;
         LAR1  #P_ADR.COMP_01;
         L     DBB[AR1, P#0.0];
         LAR1  #P_ADR.COMP_02;
         L     DIB[AR1, P#0.0];
         <>I;
         S     #AUX.DifferentValue;
         L     P#1.0;
         L     #P_ADR.COMP_01;
         +D;
         T     #P_ADR.COMP_01;
         L     P#1.0;
         L     #P_ADR.COMP_02;
         +D;
         T     #P_ADR.COMP_02;
         L     #COUNT.hA02;
         LOOP  hMP0;
         LAR1  #P_ADR.SAVE_COMP_01;
   //-------------------------------
         AN    #AUX.DifferentValue;
         JC    hB20;
         L     #LENGTH.PointerData;
         +AR1;
         L     #COUNT.hA01;
         LOOP  hA10;
         JU    hWFF;
   hWFF: NOP   0;
         L     #COUNT.hA00;
         +     1;
         T     #COUNT.hA00;
         L     #QuantityDB;
         >I;
         JC    hB40;
         JU    hA00;
   hAEE: NOP   0;
         SET;
         S     #FAULT;
         JU    END;
         JU    hAFF;
   hAFF: NOP   0;
         JU    END;
   hB20: NOP   0;
         NOP   0;
         L     #COUNT.hA00;
         JL    hB3X;
         JU    hB3X;
         JU    hB31;  //db[1]
         JU    hB32;  //db[2]
         JU    hB33;  //db[3]
         JU    hB34;  //db[4]
         JU    hB35;  //db[5]
         JU    hB36;  //db[6]
   hB3X: JU    hB3E;  //fault
   hB31: NOP   0;
         LAR1  #""Address_104";
         JU    hB3F;
   hB32: NOP   0;
         LAR1  #""Address_119";
         JU    hB3F;
   hB33: NOP   0;
         LAR1  #""Address_132";
         JU    hB3F;
   hB34: NOP   0;
         LAR1  #""Address_145";
         JU    hB3F;
   hB35: NOP   0;
         LAR1  #""Address_158";
         JU    hB3F;
   hB36: NOP   0;
         LAR1  #""Address_171";
         JU    hB3F;
   hB3E: NOP   0;
         SET;
         S     #FAULT;
         JU    END;
         JU    hB3F;
   hB3F: NOP   0;
         L     LD[AR1, P#0.0];
         T     #AUX.LD_01;
         L     LW[AR1, P#4.0];
         T     #AUX.LW_01;
         T     #PAUXnDB;
         LAR1  #""Address_464";
         L     #AUX.LD_01;
         T     LD[AR1, P#0.0];
         L     #AUX.LW_01;
         T     LW[AR1, P#4.0];
         L     #SAVE_AR1.hA10;
         T     LD[AR1, P#6.0];
         L     #P_RET_VAL.MEM;
         T     #P_RET_VAL.V[1];
         T     #P_RET_VAL.V[2];
         T     #P_RET_VAL.V[3];
         T     #P_RET_VAL.V[4];
         CALL  FILL
         ( BVAL    := #ANY_DB_DELETE,
           RET_VAL := #P_RET_VAL.V[1],
           BLK     := #Response.DeleteData
         );
         L     #P_RET_VAL.V[1];
         L     0;
         <>I;
         S     #FAULT;
         JC    END;
         CALL  FILL
         ( BVAL    := #IniData,
           RET_VAL := #P_RET_VAL.V[2],
           BLK     := #ANY_DB_DELETE
         );
         L     #P_RET_VAL.V[2];
         L     0;
         <>I;
         S     #FAULT;
         JC    END;
         S     #Response.Delete.Completed;
         L     #LogDelete;
         T     #Log.Request;
   hB3G: NOP   0;
         A     #DataInputOK;
         JC    hB3I;  //Error data input
         L     #LogDataInputNOK;
         T     #Log.Request;
   hB3I: NOP   0;
         CALL  FILL
         ( BVAL    := #DeleteData,
           RET_VAL := #P_RET_VAL.V[3],
           BLK     := #Log.DatabaseTable
         );
         L     #P_RET_VAL.V[3];
         L     0;
         <>I;
         S     #FAULT;
         JC    END;
         CALL  FILL
         ( BVAL    := #DateTime,
           RET_VAL := #P_RET_VAL.V[4],
           BLK     := #Log.DatabaseTable.DateTime
         );
         L     #P_RET_VAL.V[4];
         L     0;
         <>I;
         S     #FAULT;
         JC    END;
         JU    hB50;
   hB40: NOP   0;
         SET;
         R     #Response.Delete.Completed;
   hB50: NOP   0;
         L     #P_RET_VAL.MEM;
         T     #P_RET_VAL.V[1];
         CALL  FILL
         ( BVAL    := #DeleteData,
           RET_VAL := #P_RET_VAL.V[1],
           BLK     := #Response.Delete.BarcodeDig
         );
         L     #P_RET_VAL.V[1];
         L     0;
         <>I;
         S     #FAULT;
         JC    END;
         JU    hBFF;
   hBFF: NOP   0;
END_REGION

REGION Network 17: jA..Data input filters
         JU    jA0X;
   jA0X: NOP   0;
         JC    jAFF;
         JU    jA00;
   jA00: NOP   0;
         L     #P_RET_VAL.MEM;
         T     #NetworkReturn;
         L     #Network_17;
         T     #P_RET_VAL.MEM;
         R     #DataInputOK;
         CALL  "#DATA_INPUT_FILTER_EAN13"
         ( Data := #DigitFilter.Code.Digit,
           OK   := #DataInputOK
         );
         L     #NetworkReturn;
         L     #Network_14;
         ==I;
         JC    fAR2;  //Query
         L     #NetworkReturn;
         L     #Network_15;
         ==I;
         JC    gAR2;  //Insert
         L     #NetworkReturn;
         L     #Network_16;
         ==I;
         JC    hAR2;  //Delete
         JU    jAFF;
   jAFF: NOP   0;
END_REGION

REGION Network 18: --End--
         JU    END;
   END:  NOP   0;
         A     #FAULT;
         =     #FbFault;
         A     #DATA_ERROR;
         =     #DataError;
         L     #P_RET_VAL.MEM;
         T     #RetVal;
         LAR1  #SaveAR1;
         L     #SaveSTW;
         T     STW;
         SET;
         SAVE;
         BE;
END_REGION
END_FUNCTION_BLOCK

FUNCTION_BLOCK "#LOGGER"   // FB20, SCL
TITLE = LOGGER
{ S7_Optimized_Access := 'FALSE' }
AUTHOR : QLR
FAMILY : dnomaiD